   END_RUNG wire#w2
   RUNG wire#w1
      Contact( "DB-CompAltaDatos".Aut5 )
      Contact( "MC005-CO" )
   END_RUNG wire#w2
   RUNG wire#w1
      Contact( "DB-CompAltaDatos".Aut6 )
      Contact( "MC006-CO" )
   END_RUNG wire#w2
   RUNG wire#w1
      Contact( "DB-CompAltaDatos".TON_ParGen )
   END_RUNG wire#w2
   // the same network as SCL:
   "T_ON"(IN0 := "UNO",
          IN1 := ("DB-CompAltaDatos".Req = 0) AND (("DB-CompAltaDatos".Aut1 AND "MC001-CO") OR ("DB-CompAltaDatos".Aut2 AND "MC002-CO") OR ("DB-CompAltaDatos".Aut3 AND "MC003-CO") OR ("DB-CompAltaDatos".Aut4 AND "MC004-CO") OR ("DB-CompAltaDatos".Aut5 AND "MC005-CO") OR ("DB-CompAltaDatos".Aut6 AND "MC006-CO") OR "DB-CompAltaDatos".TON_ParGen) AND NOT "DB-CompAltaDatos".CgaPrsCrt AND NOT "DB-CompAltaDatos".PanMchCmp1 AND NOT "DB-CompAltaDatos".PanMchCmp2 AND NOT "DB-CompAltaDatos".PanMchCmp3 AND NOT "DB-CompAltaDatos".PanMchCmp4 AND NOT "DB-CompAltaDatos".PanMchCmp5,
          IN2 := "DB-CompAltaDatos".F_Osc_1seg,
          IN3 := "DB-CompAltaDatos".MinParGen,
          IO6 := "DB-CompAltaDatos".ValorParGen,
          OUT4 => "DB-CompAltaDatos".TON_ParGen,
          OUT5 => "DB-CompAltaDatos".TON_ParGen_Lim);
END_REGION

REGION Network 22
   RUNG wire#powerrail
      Contact( "DB-CompAltaDatos".TON_ParGen )
      S_SR(operand := "DB-CompAltaDatos".TON_ParGenMem, r1 := wire#w1)
   END_RUNG
   RUNG wire#powerrail
      I_Contact( "DB-CompAltaDatos".TON_ParGen )
      I_Contact( "DB-CompAltaDatos".CgaPrsCrt )
   END_RUNG wire#w1
   // the same network as SCL:
   IF "DB-CompAltaDatos".TON_ParGen THEN
       "DB-CompAltaDatos".TON_ParGenMem := TRUE;   // SR flip-flop
   END_IF;
   IF NOT "DB-CompAltaDatos".TON_ParGen AND NOT "DB-CompAltaDatos".CgaPrsCrt THEN
       "DB-CompAltaDatos".TON_ParGenMem := FALSE;
   END_IF;
END_REGION

REGION Network 23
   RUNG wire#powerrail
      Contact( "Sopladoras".Sop1 )
      S_OFFDT(T_NO := "TOFF_SP1", TV := "Sopladoras".TStopSop, R :=, BI =>, RET_VAL =>)
   END_RUNG
   // the same network as SCL:
   #_s5time1 := S_OFFDT(T_NO := "TOFF_SP1", TV := "Sopladoras".TStopSop, S := "Sopladoras".Sop1);
END_REGION

REGION Network 24
   RUNG wire#powerrail
      Contact( "Sopladoras".Sop2 )
      S_OFFDT(T_NO := "TOFF_SP2", TV := "Sopladoras".TStopSop, R :=, BI =>, RET_VAL =>)
   END_RUNG
   // the same network as SCL:
   #_s5time1 := S_OFFDT(T_NO := "TOFF_SP2", TV := "Sopladoras".TStopSop, S := "Sopladoras".Sop2);
END_REGION

REGION Network 25
   RUNG wire#powerrail
      Contact( "Sopladoras".Sop3 )
      S_OFFDT(T_NO := "TOFF_SP3", TV := "Sopladoras".TStopSop, R :=, BI =>, RET_VAL =>)
   END_RUNG
   // the same network as SCL:
   #_s5time1 := S_OFFDT(T_NO := "TOFF_SP3", TV := "Sopladoras".TStopSop, S := "Sopladoras".Sop3);
END_REGION

REGION Network 26
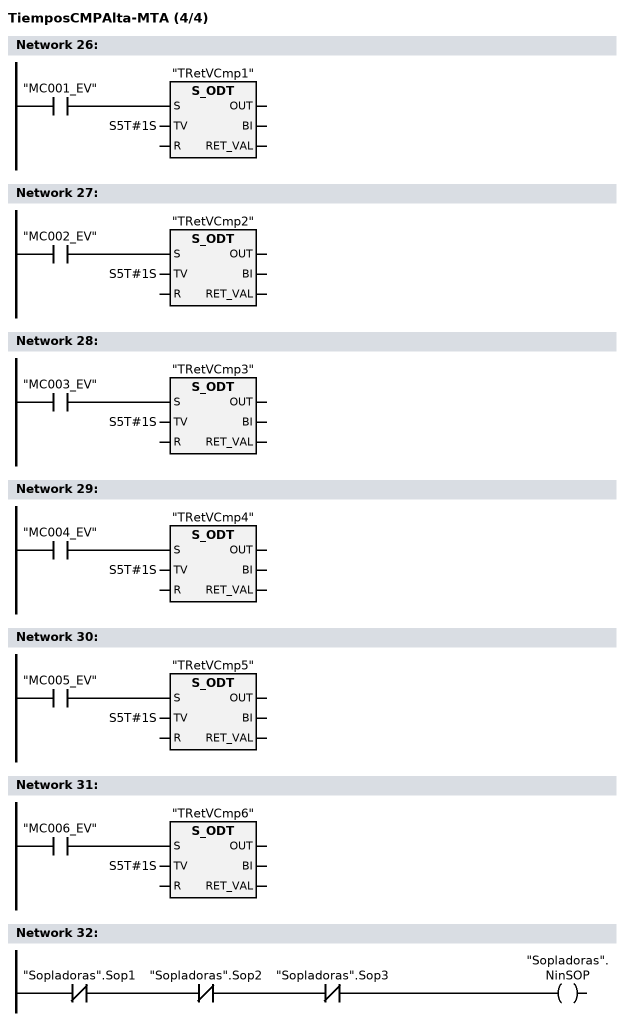
   RUNG wire#powerrail
      Contact( "MC001_EV" )
      S_ODT(T_NO := "TRetVCmp1", TV := S5T#1S, R :=, BI =>, RET_VAL =>)
   END_RUNG
   // the same network as SCL:
   #_s5time1 := S_ODT(T_NO := "TRetVCmp1", TV := S5T#1S, S := "MC001_EV");
END_REGION

REGION Network 27
   RUNG wire#powerrail
      Contact( "MC002_EV" )
      S_ODT(T_NO := "TRetVCmp2", TV := S5T#1S, R :=, BI =>, RET_VAL =>)
   END_RUNG
   // the same network as SCL:
   #_s5time1 := S_ODT(T_NO := "TRetVCmp2", TV := S5T#1S, S := "MC002_EV");
END_REGION

REGION Network 28
   RUNG wire#powerrail
      Contact( "MC003_EV" )
      S_ODT(T_NO := "TRetVCmp3", TV := S5T#1S, R :=, BI =>, RET_VAL =>)
   END_RUNG
   // the same network as SCL:
   #_s5time1 := S_ODT(T_NO := "TRetVCmp3", TV := S5T#1S, S := "MC003_EV");
END_REGION

REGION Network 29
   RUNG wire#powerrail
      Contact( "MC004_EV" )
      S_ODT(T_NO := "TRetVCmp4", TV := S5T#1S, R :=, BI =>, RET_VAL =>)
   END_RUNG
   // the same network as SCL:
   #_s5time1 := S_ODT(T_NO := "TRetVCmp4", TV := S5T#1S, S := "MC004_EV");
END_REGION

REGION Network 30
   RUNG wire#powerrail
      Contact( "MC005_EV" )
      S_ODT(T_NO := "TRetVCmp5", TV := S5T#1S, R :=, BI =>, RET_VAL =>)
   END_RUNG
   // the same network as SCL:
   #_s5time1 := S_ODT(T_NO := "TRetVCmp5", TV := S5T#1S, S := "MC005_EV");
END_REGION

REGION Network 31
   RUNG wire#powerrail
      Contact( "MC006_EV" )
      S_ODT(T_NO := "TRetVCmp6", TV := S5T#1S, R :=, BI =>, RET_VAL =>)
   END_RUNG
   // the same network as SCL:
   #_s5time1 := S_ODT(T_NO := "TRetVCmp6", S := "MC006_EV", TV := S5T#1S);
END_REGION

REGION Network 32
   RUNG wire#powerrail
      I_Contact( "Sopladoras".Sop1 )
      I_Contact( "Sopladoras".Sop2 )
      I_Contact( "Sopladoras".Sop3 )
      Coil( "Sopladoras".NinSOP )
   END_RUNG
   // the same network as SCL:
   "Sopladoras".NinSOP := NOT "Sopladoras".Sop1 AND NOT "Sopladoras".Sop2 AND NOT "Sopladoras".Sop3;
END_REGION
END_FUNCTION

FUNCTION "T_ON" : Void   // FC32, LAD
{ S7_Optimized_Access := 'FALSE' }
VERSION : 0.1
   VAR_TEMP   // added for the SCL form of the ladder/FBD networks
      _w1 : Bool;
   END_VAR
BEGIN

REGION Network 1
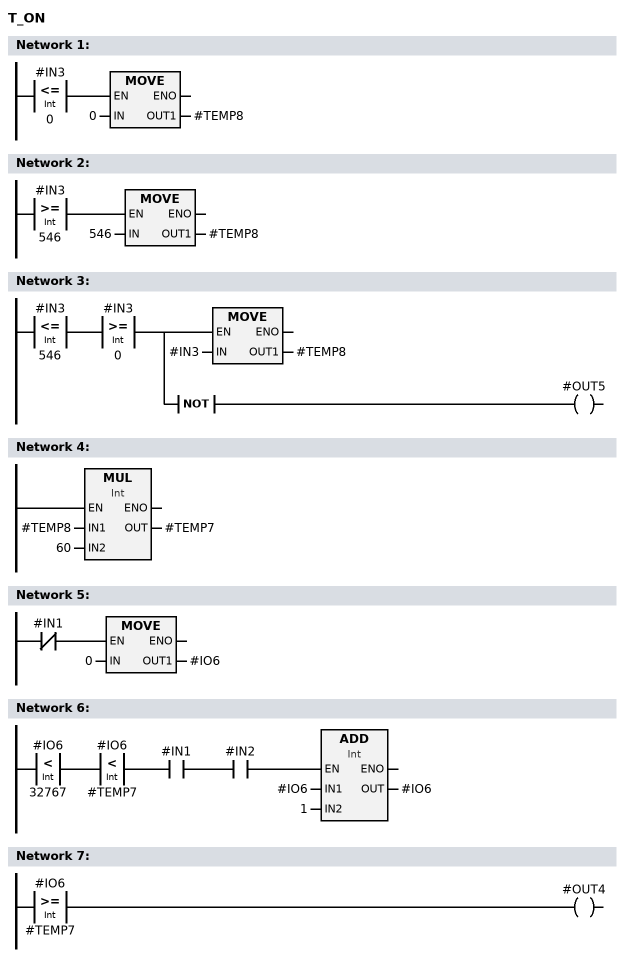
   RUNG wire#powerrail
      { S7_Templates := "SrcType := Int" } LE_Contact(in1 := #IN3, in2 := 0)
      { S7_GenerateENO := "TRUE" } Move(in := 0, out1 => #TEMP8)
   END_RUNG
   // the same network as SCL:
   IF #IN3 <= 0 THEN #TEMP8 := 0; END_IF;
END_REGION

REGION Network 2
   RUNG wire#powerrail
      { S7_Templates := "SrcType := Int" } GE_Contact(in1 := #IN3, in2 := 546)
      { S7_GenerateENO := "TRUE" } Move(in := 546, out1 => #TEMP8)
   END_RUNG
   // the same network as SCL:
   IF #IN3 >= 546 THEN #TEMP8 := 546; END_IF;
END_REGION

REGION Network 3
   RUNG wire#powerrail
      { S7_Templates := "SrcType := Int" } LE_Contact(in1 := #IN3, in2 := 546)
      { S7_Templates := "SrcType := Int" } GE_Contact(in1 := #IN3, in2 := 0)
      wire#w1
      { S7_GenerateENO := "TRUE" } Move(in := #IN3, out1 => #TEMP8)
   END_RUNG
   RUNG wire#w1
      Not()
      Coil( #OUT5 )
   END_RUNG
   // the same network as SCL:
   #_w1 := (#IN3 <= 546) AND (#IN3 >= 0);
   IF #_w1 THEN #TEMP8 := #IN3; END_IF;
   #OUT5 := NOT #_w1;
END_REGION

REGION Network 4
   RUNG wire#powerrail
      { S7_Templates := "SrcType := Int"; S7_GenerateENO := "TRUE" } Mul(in1 := #TEMP8, in2 := 60, out => #TEMP7)
   END_RUNG
   // the same network as SCL:
   #TEMP7 := #TEMP8 * 60;
END_REGION

REGION Network 5
   RUNG wire#powerrail
      I_Contact( #IN1 )
      { S7_GenerateENO := "TRUE" } Move(in := 0, out1 => #IO6)
   END_RUNG
   // the same network as SCL:
   IF NOT #IN1 THEN #IO6 := 0; END_IF;
END_REGION

REGION Network 6
   RUNG wire#powerrail
      { S7_Templates := "SrcType := Int" } LT_Contact(in1 := #IO6, in2 := 32767)
      { S7_Templates := "SrcType := Int" } LT_Contact(in1 := #IO6, in2 := #TEMP7)
      Contact( #IN1 )
      Contact( #IN2 )
      { S7_Templates := "SrcType := Int"; S7_GenerateENO := "TRUE" } Add(in1 := #IO6, in2 := 1, out => #IO6)
   END_RUNG
   // the same network as SCL:
   IF (#IO6 < 32767) AND (#IO6 < #TEMP7) AND #IN1 AND #IN2 THEN #IO6 := #IO6 + 1; END_IF;
END_REGION

REGION Network 7
   RUNG wire#powerrail
      { S7_Templates := "SrcType := Int" } GE_Contact(in1 := #IO6, in2 := #TEMP7)
      Coil( #OUT4 )
   END_RUNG
   // the same network as SCL:
   #OUT4 := #IO6 >= #TEMP7;
END_REGION
END_FUNCTION

FUNCTION "PrioridadesCmpAlta" : Void   // FC33, LAD
{ S7_Optimized_Access := 'FALSE' }
VERSION : 0.1
   VAR_TEMP   // added for the SCL form of the ladder/FBD networks
      _w1 : Bool;
   END_VAR
BEGIN

REGION Network 1
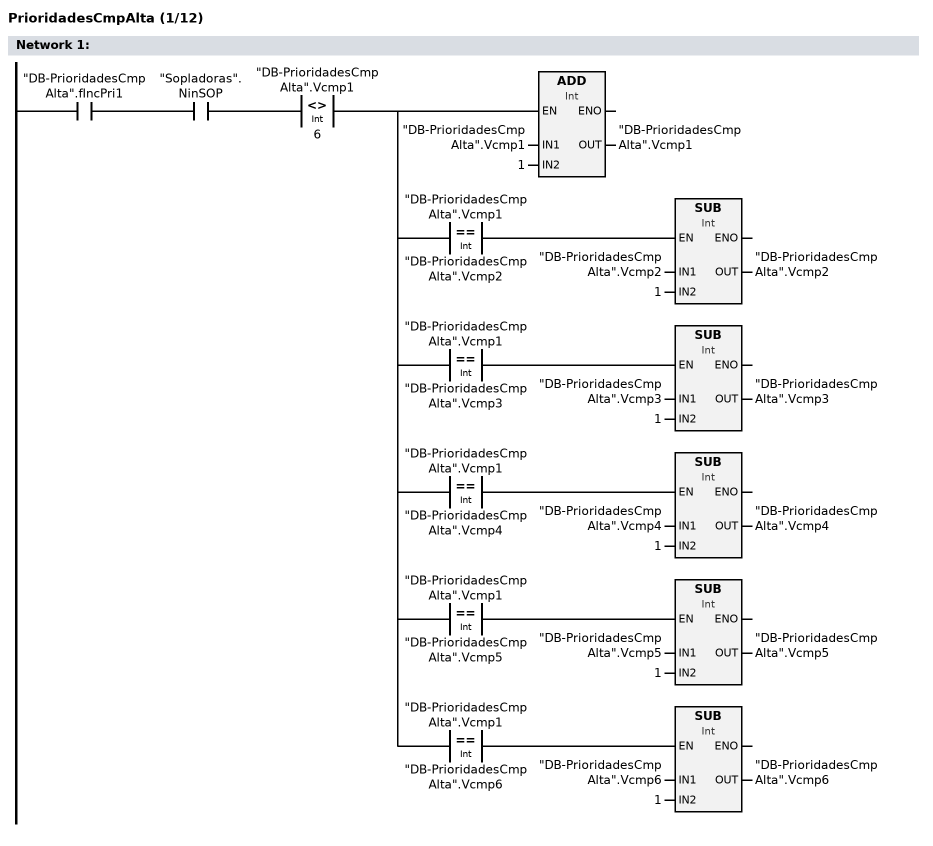
   RUNG wire#powerrail
      Contact( "DB-PrioridadesCmpAlta".fIncPri1 )
      Contact( "Sopladoras".NinSOP )
      { S7_Templates := "SrcType := Int" } NE_Contact(in1 := "DB-PrioridadesCmpAlta".Vcmp1, in2 := 6)
      wire#w1
      { S7_Templates := "SrcType := Int"; S7_GenerateENO := "TRUE" } Add(in1 := "DB-PrioridadesCmpAlta".Vcmp1, in2 := 1, out => "DB-PrioridadesCmpAlta".Vcmp1)
   END_RUNG
   RUNG wire#w1
      { S7_Templates := "SrcType := Int" } EQ_Contact(in1 := "DB-PrioridadesCmpAlta".Vcmp1, in2 := "DB-PrioridadesCmpAlta".Vcmp2)
      { S7_Templates := "SrcType := Int"; S7_GenerateENO := "TRUE" } Sub(in1 := "DB-PrioridadesCmpAlta".Vcmp2, in2 := 1, out => "DB-PrioridadesCmpAlta".Vcmp2)
   END_RUNG
   RUNG wire#w1
      { S7_Templates := "SrcType := Int" } EQ_Contact(in1 := "DB-PrioridadesCmpAlta".Vcmp1, in2 := "DB-PrioridadesCmpAlta".Vcmp3)
      { S7_Templates := "SrcType := Int"; S7_GenerateENO := "TRUE" } Sub(in1 := "DB-PrioridadesCmpAlta".Vcmp3, in2 := 1, out => "DB-PrioridadesCmpAlta".Vcmp3)
   END_RUNG
   RUNG wire#w1
      { S7_Templates := "SrcType := Int" } EQ_Contact(in1 := "DB-PrioridadesCmpAlta".Vcmp1, in2 := "DB-PrioridadesCmpAlta".Vcmp4)
      { S7_Templates := "SrcType := Int"; S7_GenerateENO := "TRUE" } Sub(in1 := "DB-PrioridadesCmpAlta".Vcmp4, in2 := 1, out => "DB-PrioridadesCmpAlta".Vcmp4)
   END_RUNG
   RUNG wire#w1
      { S7_Templates := "SrcType := Int" } EQ_Contact(in1 := "DB-PrioridadesCmpAlta".Vcmp1, in2 := "DB-PrioridadesCmpAlta".Vcmp5)
      { S7_Templates := "SrcType := Int"; S7_GenerateENO := "TRUE" } Sub(in1 := "DB-PrioridadesCmpAlta".Vcmp5, in2 := 1, out => "DB-PrioridadesCmpAlta".Vcmp5)
   END_RUNG
   RUNG wire#w1
      { S7_Templates := "SrcType := Int" } EQ_Contact(in1 := "DB-PrioridadesCmpAlta".Vcmp1, in2 := "DB-PrioridadesCmpAlta".Vcmp6)
      { S7_Templates := "SrcType := Int"; S7_GenerateENO := "TRUE" } Sub(in1 := "DB-PrioridadesCmpAlta".Vcmp6, in2 := 1, out => "DB-PrioridadesCmpAlta".Vcmp6)
   END_RUNG
   // the same network as SCL:
   #_w1 := "DB-PrioridadesCmpAlta".fIncPri1 AND "Sopladoras".NinSOP AND ("DB-PrioridadesCmpAlta".Vcmp1 <> 6);
   IF #_w1 THEN "DB-PrioridadesCmpAlta".Vcmp1 := "DB-PrioridadesCmpAlta".Vcmp1 + 1; END_IF;
   IF #_w1 AND ("DB-PrioridadesCmpAlta".Vcmp1 = "DB-PrioridadesCmpAlta".Vcmp2) THEN
       "DB-PrioridadesCmpAlta".Vcmp2 := "DB-PrioridadesCmpAlta".Vcmp2 - 1;
   END_IF;
   IF #_w1 AND ("DB-PrioridadesCmpAlta".Vcmp1 = "DB-PrioridadesCmpAlta".Vcmp3) THEN
       "DB-PrioridadesCmpAlta".Vcmp3 := "DB-PrioridadesCmpAlta".Vcmp3 - 1;
   END_IF;
   IF #_w1 AND ("DB-PrioridadesCmpAlta".Vcmp1 = "DB-PrioridadesCmpAlta".Vcmp4) THEN
       "DB-PrioridadesCmpAlta".Vcmp4 := "DB-PrioridadesCmpAlta".Vcmp4 - 1;
   END_IF;
   IF #_w1 AND ("DB-PrioridadesCmpAlta".Vcmp1 = "DB-PrioridadesCmpAlta".Vcmp5) THEN
       "DB-PrioridadesCmpAlta".Vcmp5 := "DB-PrioridadesCmpAlta".Vcmp5 - 1;
   END_IF;
   IF #_w1 AND ("DB-PrioridadesCmpAlta".Vcmp1 = "DB-PrioridadesCmpAlta".Vcmp6) THEN
       "DB-PrioridadesCmpAlta".Vcmp6 := "DB-PrioridadesCmpAlta".Vcmp6 - 1;
   END_IF;
END_REGION

REGION Network 2
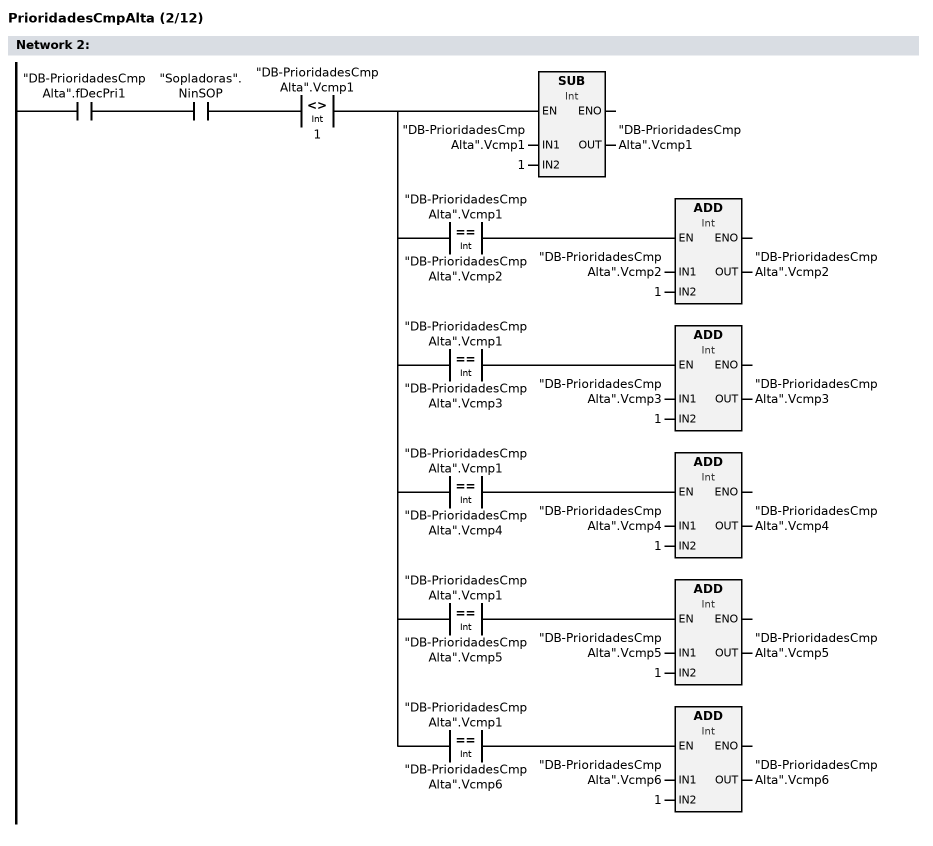
   RUNG wire#powerrail
      Contact( "DB-PrioridadesCmpAlta".fDecPri1 )
      Contact( "Sopladoras".NinSOP )
      { S7_Templates := "SrcType := Int" } NE_Contact(in1 := "DB-PrioridadesCmpAlta".Vcmp1, in2 := 1)
      wire#w1
      { S7_Templates := "SrcType := Int"; S7_GenerateENO := "TRUE" } Sub(in1 := "DB-PrioridadesCmpAlta".Vcmp1, in2 := 1, out => "DB-PrioridadesCmpAlta".Vcmp1)
   END_RUNG
   RUNG wire#w1
      { S7_Templates := "SrcType := Int" } EQ_Contact(in1 := "DB-PrioridadesCmpAlta".Vcmp1, in2 := "DB-PrioridadesCmpAlta".Vcmp2)
      { S7_Templates := "SrcType := Int"; S7_GenerateENO := "TRUE" } Add(in1 := "DB-PrioridadesCmpAlta".Vcmp2, in2 := 1, out => "DB-PrioridadesCmpAlta".Vcmp2)
   END_RUNG
   RUNG wire#w1
      { S7_Templates := "SrcType := Int" } EQ_Contact(in1 := "DB-PrioridadesCmpAlta".Vcmp1, in2 := "DB-PrioridadesCmpAlta".Vcmp3)
      { S7_Templates := "SrcType := Int"; S7_GenerateENO := "TRUE" } Add(in1 := "DB-PrioridadesCmpAlta".Vcmp3, in2 := 1, out => "DB-PrioridadesCmpAlta".Vcmp3)
   END_RUNG
   RUNG wire#w1
      { S7_Templates := "SrcType := Int" } EQ_Contact(in1 := "DB-PrioridadesCmpAlta".Vcmp1, in2 := "DB-PrioridadesCmpAlta".Vcmp4)
      { S7_Templates := "SrcType := Int"; S7_GenerateENO := "TRUE" } Add(in1 := "DB-PrioridadesCmpAlta".Vcmp4, in2 := 1, out => "DB-PrioridadesCmpAlta".Vcmp4)
   END_RUNG
   RUNG wire#w1
      { S7_Templates := "SrcType := Int" } EQ_Contact(in1 := "DB-PrioridadesCmpAlta".Vcmp1, in2 := "DB-PrioridadesCmpAlta".Vcmp5)
      { S7_Templates := "SrcType := Int"; S7_GenerateENO := "TRUE" } Add(in1 := "DB-PrioridadesCmpAlta".Vcmp5, in2 := 1, out => "DB-PrioridadesCmpAlta".Vcmp5)
   END_RUNG
   RUNG wire#w1
      { S7_Templates := "SrcType := Int" } EQ_Contact(in1 := "DB-PrioridadesCmpAlta".Vcmp1, in2 := "DB-PrioridadesCmpAlta".Vcmp6)
      { S7_Templates := "SrcType := Int"; S7_GenerateENO := "TRUE" } Add(in1 := "DB-PrioridadesCmpAlta".Vcmp6, in2 := 1, out => "DB-PrioridadesCmpAlta".Vcmp6)
   END_RUNG
   // the same network as SCL:
   #_w1 := "DB-PrioridadesCmpAlta".fDecPri1 AND "Sopladoras".NinSOP AND ("DB-PrioridadesCmpAlta".Vcmp1 <> 1);
   IF #_w1 THEN "DB-PrioridadesCmpAlta".Vcmp1 := "DB-PrioridadesCmpAlta".Vcmp1 - 1; END_IF;
   IF #_w1 AND ("DB-PrioridadesCmpAlta".Vcmp1 = "DB-PrioridadesCmpAlta".Vcmp2) THEN
       "DB-PrioridadesCmpAlta".Vcmp2 := "DB-PrioridadesCmpAlta".Vcmp2 + 1;
   END_IF;
   IF #_w1 AND ("DB-PrioridadesCmpAlta".Vcmp1 = "DB-PrioridadesCmpAlta".Vcmp3) THEN
       "DB-PrioridadesCmpAlta".Vcmp3 := "DB-PrioridadesCmpAlta".Vcmp3 + 1;
   END_IF;
   IF #_w1 AND ("DB-PrioridadesCmpAlta".Vcmp1 = "DB-PrioridadesCmpAlta".Vcmp4) THEN
       "DB-PrioridadesCmpAlta".Vcmp4 := "DB-PrioridadesCmpAlta".Vcmp4 + 1;
   END_IF;
   IF #_w1 AND ("DB-PrioridadesCmpAlta".Vcmp1 = "DB-PrioridadesCmpAlta".Vcmp5) THEN
       "DB-PrioridadesCmpAlta".Vcmp5 := "DB-PrioridadesCmpAlta".Vcmp5 + 1;
   END_IF;
   IF #_w1 AND ("DB-PrioridadesCmpAlta".Vcmp1 = "DB-PrioridadesCmpAlta".Vcmp6) THEN
       "DB-PrioridadesCmpAlta".Vcmp6 := "DB-PrioridadesCmpAlta".Vcmp6 + 1;
   END_IF;
END_REGION

REGION Network 3
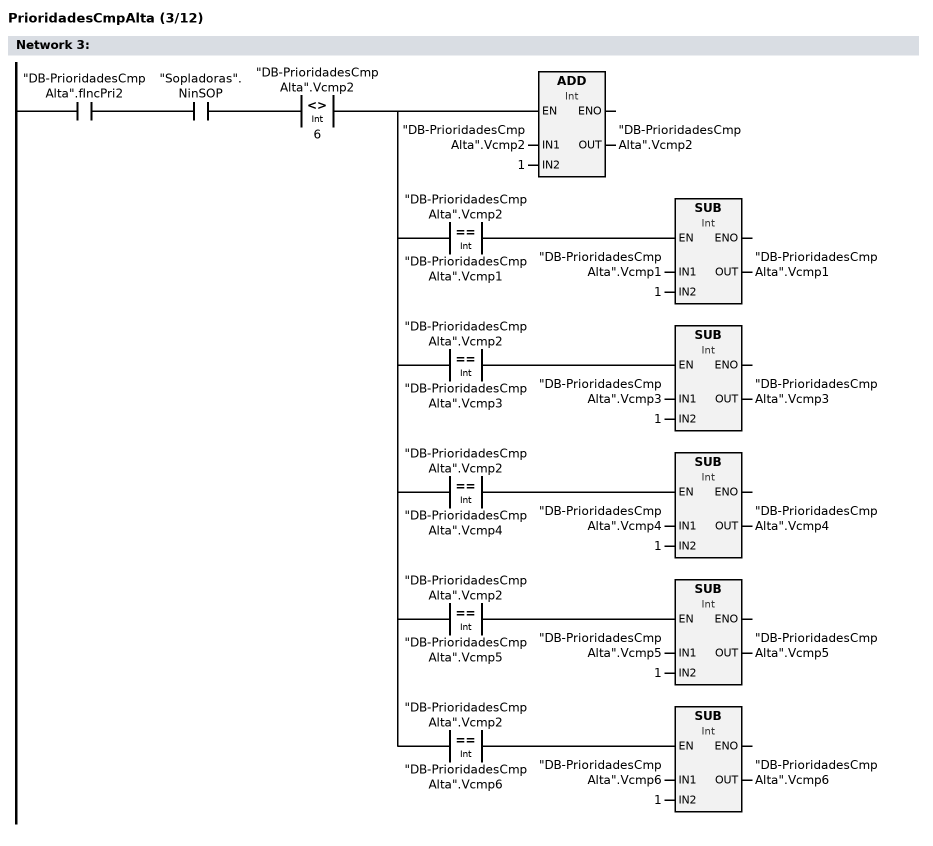
   RUNG wire#powerrail
      Contact( "DB-PrioridadesCmpAlta".fIncPri2 )
      Contact( "Sopladoras".NinSOP )
      { S7_Templates := "SrcType := Int" } NE_Contact(in1 := "DB-PrioridadesCmpAlta".Vcmp2, in2 := 6)
      wire#w1
      { S7_Templates := "SrcType := Int"; S7_GenerateENO := "TRUE" } Add(in1 := "DB-PrioridadesCmpAlta".Vcmp2, in2 := 1, out => "DB-PrioridadesCmpAlta".Vcmp2)
   END_RUNG
   RUNG wire#w1
      { S7_Templates := "SrcType := Int" } EQ_Contact(in1 := "DB-PrioridadesCmpAlta".Vcmp2, in2 := "DB-PrioridadesCmpAlta".Vcmp1)
      { S7_Templates := "SrcType := Int"; S7_GenerateENO := "TRUE" } Sub(in1 := "DB-PrioridadesCmpAlta".Vcmp1, in2 := 1, out => "DB-PrioridadesCmpAlta".Vcmp1)
   END_RUNG
   RUNG wire#w1
      { S7_Templates := "SrcType := Int" } EQ_Contact(in1 := "DB-PrioridadesCmpAlta".Vcmp2, in2 := "DB-PrioridadesCmpAlta".Vcmp3)
      { S7_Templates := "SrcType := Int"; S7_GenerateENO := "TRUE" } Sub(in1 := "DB-PrioridadesCmpAlta".Vcmp3, in2 := 1, out => "DB-PrioridadesCmpAlta".Vcmp3)
   END_RUNG
   RUNG wire#w1
      { S7_Templates := "SrcType := Int" } EQ_Contact(in1 := "DB-PrioridadesCmpAlta".Vcmp2, in2 := "DB-PrioridadesCmpAlta".Vcmp4)
      { S7_Templates := "SrcType := Int"; S7_GenerateENO := "TRUE" } Sub(in1 := "DB-PrioridadesCmpAlta".Vcmp4, in2 := 1, out => "DB-PrioridadesCmpAlta".Vcmp4)
   END_RUNG
   RUNG wire#w1
      { S7_Templates := "SrcType := Int" } EQ_Contact(in1 := "DB-PrioridadesCmpAlta".Vcmp2, in2 := "DB-PrioridadesCmpAlta".Vcmp5)
      { S7_Templates := "SrcType := Int"; S7_GenerateENO := "TRUE" } Sub(in1 := "DB-PrioridadesCmpAlta".Vcmp5, in2 := 1, out => "DB-PrioridadesCmpAlta".Vcmp5)
   END_RUNG
   RUNG wire#w1
      { S7_Templates := "SrcType := Int" } EQ_Contact(in1 := "DB-PrioridadesCmpAlta".Vcmp2, in2 := "DB-PrioridadesCmpAlta".Vcmp6)
      { S7_Templates := "SrcType := Int"; S7_GenerateENO := "TRUE" } Sub(in1 := "DB-PrioridadesCmpAlta".Vcmp6, in2 := 1, out => "DB-PrioridadesCmpAlta".Vcmp6)
   END_RUNG
   // the same network as SCL:
   #_w1 := "DB-PrioridadesCmpAlta".fIncPri2 AND "Sopladoras".NinSOP AND ("DB-PrioridadesCmpAlta".Vcmp2 <> 6);
   IF #_w1 THEN "DB-PrioridadesCmpAlta".Vcmp2 := "DB-PrioridadesCmpAlta".Vcmp2 + 1; END_IF;
   IF #_w1 AND ("DB-PrioridadesCmpAlta".Vcmp2 = "DB-PrioridadesCmpAlta".Vcmp1) THEN
       "DB-PrioridadesCmpAlta".Vcmp1 := "DB-PrioridadesCmpAlta".Vcmp1 - 1;
   END_IF;
   IF #_w1 AND ("DB-PrioridadesCmpAlta".Vcmp2 = "DB-PrioridadesCmpAlta".Vcmp3) THEN
       "DB-PrioridadesCmpAlta".Vcmp3 := "DB-PrioridadesCmpAlta".Vcmp3 - 1;
   END_IF;
   IF #_w1 AND ("DB-PrioridadesCmpAlta".Vcmp2 = "DB-PrioridadesCmpAlta".Vcmp4) THEN
       "DB-PrioridadesCmpAlta".Vcmp4 := "DB-PrioridadesCmpAlta".Vcmp4 - 1;
   END_IF;
   IF #_w1 AND ("DB-PrioridadesCmpAlta".Vcmp2 = "DB-PrioridadesCmpAlta".Vcmp5) THEN
       "DB-PrioridadesCmpAlta".Vcmp5 := "DB-PrioridadesCmpAlta".Vcmp5 - 1;
   END_IF;
   IF #_w1 AND ("DB-PrioridadesCmpAlta".Vcmp2 = "DB-PrioridadesCmpAlta".Vcmp6) THEN
       "DB-PrioridadesCmpAlta".Vcmp6 := "DB-PrioridadesCmpAlta".Vcmp6 - 1;
   END_IF;
END_REGION

REGION Network 4
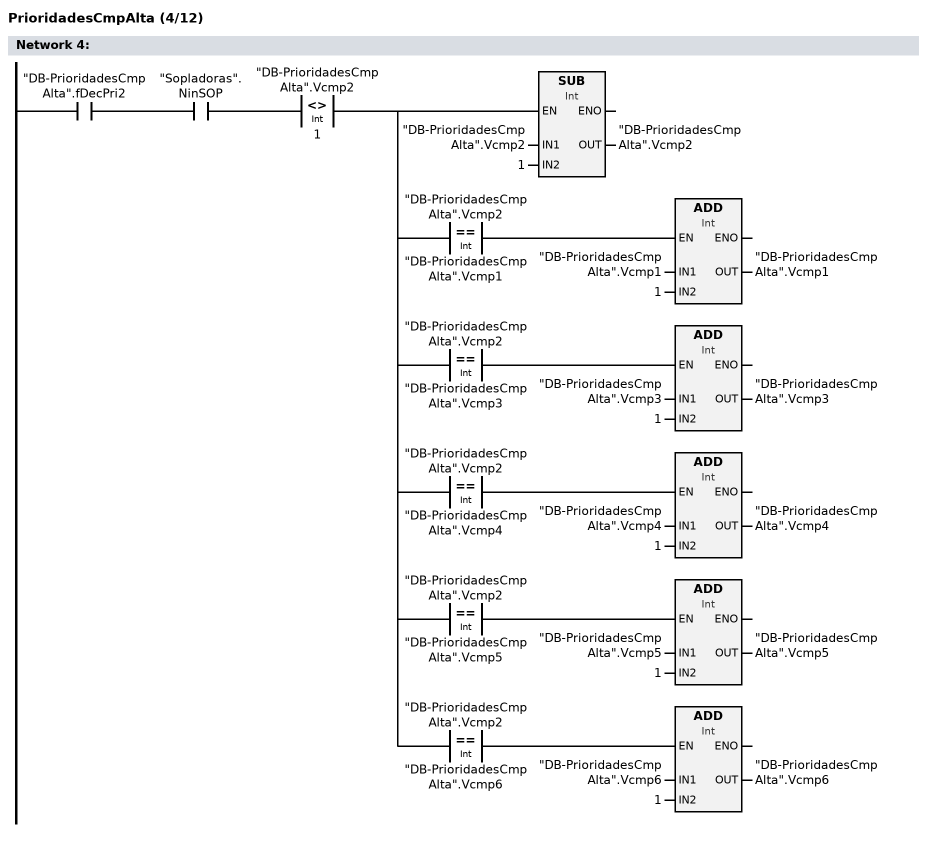
   RUNG wire#powerrail
      Contact( "DB-PrioridadesCmpAlta".fDecPri2 )
      Contact( "Sopladoras".NinSOP )
      { S7_Templates := "SrcType := Int" } NE_Contact(in1 := "DB-PrioridadesCmpAlta".Vcmp2, in2 := 1)
      wire#w1
      { S7_Templates := "SrcType := Int"; S7_GenerateENO := "TRUE" } Sub(in1 := "DB-PrioridadesCmpAlta".Vcmp2, in2 := 1, out => "DB-PrioridadesCmpAlta".Vcmp2)
   END_RUNG
   RUNG wire#w1
      { S7_Templates := "SrcType := Int" } EQ_Contact(in1 := "DB-PrioridadesCmpAlta".Vcmp2, in2 := "DB-PrioridadesCmpAlta".Vcmp1)
      { S7_Templates := "SrcType := Int"; S7_GenerateENO := "TRUE" } Add(in1 := "DB-PrioridadesCmpAlta".Vcmp1, in2 := 1, out => "DB-PrioridadesCmpAlta".Vcmp1)
   END_RUNG
   RUNG wire#w1
      { S7_Templates := "SrcType := Int" } EQ_Contact(in1 := "DB-PrioridadesCmpAlta".Vcmp2, in2 := "DB-PrioridadesCmpAlta".Vcmp3)
      { S7_Templates := "SrcType := Int"; S7_GenerateENO := "TRUE" } Add(in1 := "DB-PrioridadesCmpAlta".Vcmp3, in2 := 1, out => "DB-PrioridadesCmpAlta".Vcmp3)
   END_RUNG
   RUNG wire#w1
      { S7_Templates := "SrcType := Int" } EQ_Contact(in1 := "DB-PrioridadesCmpAlta".Vcmp2, in2 := "DB-PrioridadesCmpAlta".Vcmp4)
      { S7_Templates := "SrcType := Int"; S7_GenerateENO := "TRUE" } Add(in1 := "DB-PrioridadesCmpAlta".Vcmp4, in2 := 1, out => "DB-PrioridadesCmpAlta".Vcmp4)
   END_RUNG
   RUNG wire#w1
      { S7_Templates := "SrcType := Int" } EQ_Contact(in1 := "DB-PrioridadesCmpAlta".Vcmp2, in2 := "DB-PrioridadesCmpAlta".Vcmp5)
      { S7_Templates := "SrcType := Int"; S7_GenerateENO := "TRUE" } Add(in1 := "DB-PrioridadesCmpAlta".Vcmp5, in2 := 1, out => "DB-PrioridadesCmpAlta".Vcmp5)
   END_RUNG
   RUNG wire#w1
      { S7_Templates := "SrcType := Int" } EQ_Contact(in1 := "DB-PrioridadesCmpAlta".Vcmp2, in2 := "DB-PrioridadesCmpAlta".Vcmp6)
      { S7_Templates := "SrcType := Int"; S7_GenerateENO := "TRUE" } Add(in1 := "DB-PrioridadesCmpAlta".Vcmp6, in2 := 1, out => "DB-PrioridadesCmpAlta".Vcmp6)
   END_RUNG
   // the same network as SCL:
   #_w1 := "DB-PrioridadesCmpAlta".fDecPri2 AND "Sopladoras".NinSOP AND ("DB-PrioridadesCmpAlta".Vcmp2 <> 1);
   IF #_w1 THEN "DB-PrioridadesCmpAlta".Vcmp2 := "DB-PrioridadesCmpAlta".Vcmp2 - 1; END_IF;
   IF #_w1 AND ("DB-PrioridadesCmpAlta".Vcmp2 = "DB-PrioridadesCmpAlta".Vcmp1) THEN
       "DB-PrioridadesCmpAlta".Vcmp1 := "DB-PrioridadesCmpAlta".Vcmp1 + 1;
   END_IF;
   IF #_w1 AND ("DB-PrioridadesCmpAlta".Vcmp2 = "DB-PrioridadesCmpAlta".Vcmp3) THEN
       "DB-PrioridadesCmpAlta".Vcmp3 := "DB-PrioridadesCmpAlta".Vcmp3 + 1;
   END_IF;
   IF #_w1 AND ("DB-PrioridadesCmpAlta".Vcmp2 = "DB-PrioridadesCmpAlta".Vcmp4) THEN
       "DB-PrioridadesCmpAlta".Vcmp4 := "DB-PrioridadesCmpAlta".Vcmp4 + 1;
   END_IF;
   IF #_w1 AND ("DB-PrioridadesCmpAlta".Vcmp2 = "DB-PrioridadesCmpAlta".Vcmp5) THEN
       "DB-PrioridadesCmpAlta".Vcmp5 := "DB-PrioridadesCmpAlta".Vcmp5 + 1;
   END_IF;
   IF #_w1 AND ("DB-PrioridadesCmpAlta".Vcmp2 = "DB-PrioridadesCmpAlta".Vcmp6) THEN
       "DB-PrioridadesCmpAlta".Vcmp6 := "DB-PrioridadesCmpAlta".Vcmp6 + 1;
   END_IF;
END_REGION

REGION Network 5
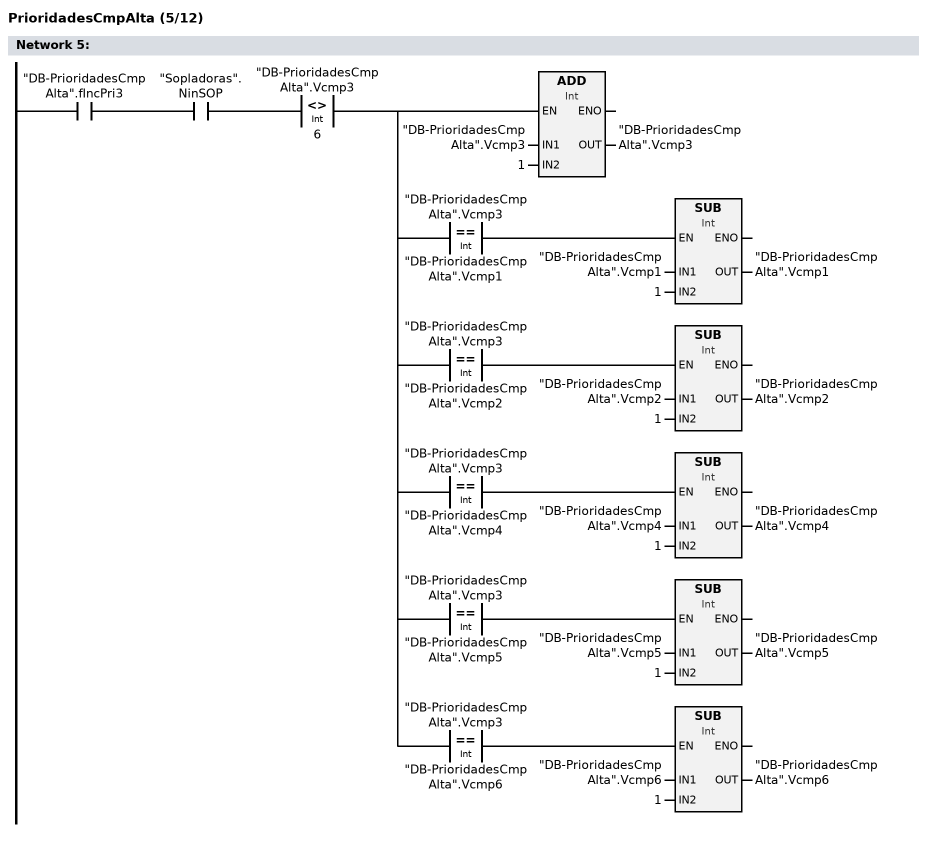
   RUNG wire#powerrail
      Contact( "DB-PrioridadesCmpAlta".fIncPri3 )
      Contact( "Sopladoras".NinSOP )
      { S7_Templates := "SrcType := Int" } NE_Contact(in1 := "DB-PrioridadesCmpAlta".Vcmp3, in2 := 6)
      wire#w1
      { S7_Templates := "SrcType := Int"; S7_GenerateENO := "TRUE" } Add(in1 := "DB-PrioridadesCmpAlta".Vcmp3, in2 := 1, out => "DB-PrioridadesCmpAlta".Vcmp3)
   END_RUNG
   RUNG wire#w1
      { S7_Templates := "SrcType := Int" } EQ_Contact(in1 := "DB-PrioridadesCmpAlta".Vcmp3, in2 := "DB-PrioridadesCmpAlta".Vcmp1)
      { S7_Templates := "SrcType := Int"; S7_GenerateENO := "TRUE" } Sub(in1 := "DB-PrioridadesCmpAlta".Vcmp1, in2 := 1, out => "DB-PrioridadesCmpAlta".Vcmp1)
   END_RUNG
   RUNG wire#w1
      { S7_Templates := "SrcType := Int" } EQ_Contact(in1 := "DB-PrioridadesCmpAlta".Vcmp3, in2 := "DB-PrioridadesCmpAlta".Vcmp2)
      { S7_Templates := "SrcType := Int"; S7_GenerateENO := "TRUE" } Sub(in1 := "DB-PrioridadesCmpAlta".Vcmp2, in2 := 1, out => "DB-PrioridadesCmpAlta".Vcmp2)
   END_RUNG
   RUNG wire#w1
      { S7_Templates := "SrcType := Int" } EQ_Contact(in1 := "DB-PrioridadesCmpAlta".Vcmp3, in2 := "DB-PrioridadesCmpAlta".Vcmp4)
      { S7_Templates := "SrcType := Int"; S7_GenerateENO := "TRUE" } Sub(in1 := "DB-PrioridadesCmpAlta".Vcmp4, in2 := 1, out => "DB-PrioridadesCmpAlta".Vcmp4)
   END_RUNG
   RUNG wire#w1
      { S7_Templates := "SrcType := Int" } EQ_Contact(in1 := "DB-PrioridadesCmpAlta".Vcmp3, in2 := "DB-PrioridadesCmpAlta".Vcmp5)
      { S7_Templates := "SrcType := Int"; S7_GenerateENO := "TRUE" } Sub(in1 := "DB-PrioridadesCmpAlta".Vcmp5, in2 := 1, out => "DB-PrioridadesCmpAlta".Vcmp5)
   END_RUNG
   RUNG wire#w1
      { S7_Templates := "SrcType := Int" } EQ_Contact(in1 := "DB-PrioridadesCmpAlta".Vcmp3, in2 := "DB-PrioridadesCmpAlta".Vcmp6)
      { S7_Templates := "SrcType := Int"; S7_GenerateENO := "TRUE" } Sub(in1 := "DB-PrioridadesCmpAlta".Vcmp6, in2 := 1, out => "DB-PrioridadesCmpAlta".Vcmp6)
   END_RUNG
   // the same network as SCL:
   #_w1 := "DB-PrioridadesCmpAlta".fIncPri3 AND "Sopladoras".NinSOP AND ("DB-PrioridadesCmpAlta".Vcmp3 <> 6);
   IF #_w1 THEN "DB-PrioridadesCmpAlta".Vcmp3 := "DB-PrioridadesCmpAlta".Vcmp3 + 1; END_IF;
   IF #_w1 AND ("DB-PrioridadesCmpAlta".Vcmp3 = "DB-PrioridadesCmpAlta".Vcmp1) THEN
       "DB-PrioridadesCmpAlta".Vcmp1 := "DB-PrioridadesCmpAlta".Vcmp1 - 1;
   END_IF;
   IF #_w1 AND ("DB-PrioridadesCmpAlta".Vcmp3 = "DB-PrioridadesCmpAlta".Vcmp2) THEN
       "DB-PrioridadesCmpAlta".Vcmp2 := "DB-PrioridadesCmpAlta".Vcmp2 - 1;
   END_IF;
   IF #_w1 AND ("DB-PrioridadesCmpAlta".Vcmp3 = "DB-PrioridadesCmpAlta".Vcmp4) THEN
       "DB-PrioridadesCmpAlta".Vcmp4 := "DB-PrioridadesCmpAlta".Vcmp4 - 1;
   END_IF;
   IF #_w1 AND ("DB-PrioridadesCmpAlta".Vcmp3 = "DB-PrioridadesCmpAlta".Vcmp5) THEN
       "DB-PrioridadesCmpAlta".Vcmp5 := "DB-PrioridadesCmpAlta".Vcmp5 - 1;
   END_IF;
   IF #_w1 AND ("DB-PrioridadesCmpAlta".Vcmp3 = "DB-PrioridadesCmpAlta".Vcmp6) THEN
       "DB-PrioridadesCmpAlta".Vcmp6 := "DB-PrioridadesCmpAlta".Vcmp6 - 1;
   END_IF;
END_REGION

REGION Network 6
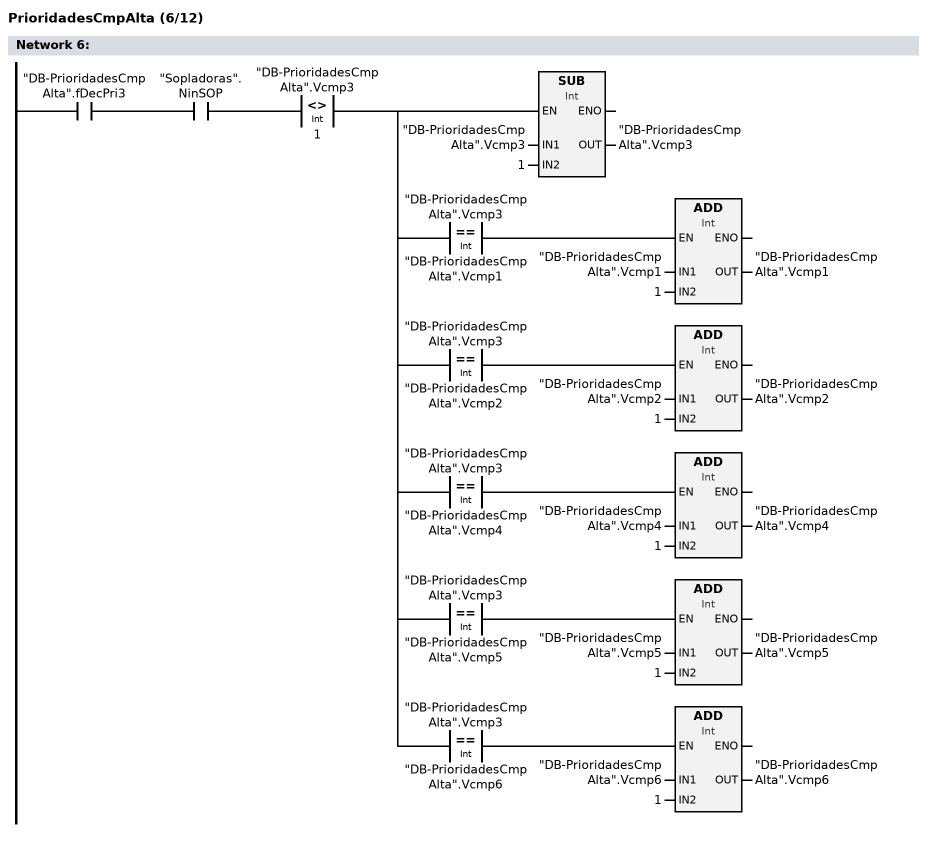
   RUNG wire#powerrail
      Contact( "DB-PrioridadesCmpAlta".fDecPri3 )
      Contact( "Sopladoras".NinSOP )
      { S7_Templates := "SrcType := Int" } NE_Contact(in1 := "DB-PrioridadesCmpAlta".Vcmp3, in2 := 1)
      wire#w1
      { S7_Templates := "SrcType := Int"; S7_GenerateENO := "TRUE" } Sub(in1 := "DB-PrioridadesCmpAlta".Vcmp3, in2 := 1, out => "DB-PrioridadesCmpAlta".Vcmp3)
   END_RUNG
   RUNG wire#w1
      { S7_Templates := "SrcType := Int" } EQ_Contact(in1 := "DB-PrioridadesCmpAlta".Vcmp3, in2 := "DB-PrioridadesCmpAlta".Vcmp1)
      { S7_Templates := "SrcType := Int"; S7_GenerateENO := "TRUE" } Add(in1 := "DB-PrioridadesCmpAlta".Vcmp1, in2 := 1, out => "DB-PrioridadesCmpAlta".Vcmp1)
   END_RUNG
   RUNG wire#w1
      { S7_Templates := "SrcType := Int" } EQ_Contact(in1 := "DB-PrioridadesCmpAlta".Vcmp3, in2 := "DB-PrioridadesCmpAlta".Vcmp2)
      { S7_Templates := "SrcType := Int"; S7_GenerateENO := "TRUE" } Add(in1 := "DB-PrioridadesCmpAlta".Vcmp2, in2 := 1, out => "DB-PrioridadesCmpAlta".Vcmp2)
   END_RUNG
   RUNG wire#w1
      { S7_Templates := "SrcType := Int" } EQ_Contact(in1 := "DB-PrioridadesCmpAlta".Vcmp3, in2 := "DB-PrioridadesCmpAlta".Vcmp4)
      { S7_Templates := "SrcType := Int"; S7_GenerateENO := "TRUE" } Add(in1 := "DB-PrioridadesCmpAlta".Vcmp4, in2 := 1, out => "DB-PrioridadesCmpAlta".Vcmp4)
   END_RUNG
   RUNG wire#w1
      { S7_Templates := "SrcType := Int" } EQ_Contact(in1 := "DB-PrioridadesCmpAlta".Vcmp3, in2 := "DB-PrioridadesCmpAlta".Vcmp5)
      { S7_Templates := "SrcType := Int"; S7_GenerateENO := "TRUE" } Add(in1 := "DB-PrioridadesCmpAlta".Vcmp5, in2 := 1, out => "DB-PrioridadesCmpAlta".Vcmp5)
   END_RUNG
   RUNG wire#w1
      { S7_Templates := "SrcType := Int" } EQ_Contact(in1 := "DB-PrioridadesCmpAlta".Vcmp3, in2 := "DB-PrioridadesCmpAlta".Vcmp6)
      { S7_Templates := "SrcType := Int"; S7_GenerateENO := "TRUE" } Add(in1 := "DB-PrioridadesCmpAlta".Vcmp6, in2 := 1, out => "DB-PrioridadesCmpAlta".Vcmp6)
   END_RUNG
   // the same network as SCL:
   #_w1 := "DB-PrioridadesCmpAlta".fDecPri3 AND "Sopladoras".NinSOP AND ("DB-PrioridadesCmpAlta".Vcmp3 <> 1);
   IF #_w1 THEN "DB-PrioridadesCmpAlta".Vcmp3 := "DB-PrioridadesCmpAlta".Vcmp3 - 1; END_IF;
   IF #_w1 AND ("DB-PrioridadesCmpAlta".Vcmp3 = "DB-PrioridadesCmpAlta".Vcmp1) THEN
       "DB-PrioridadesCmpAlta".Vcmp1 := "DB-PrioridadesCmpAlta".Vcmp1 + 1;